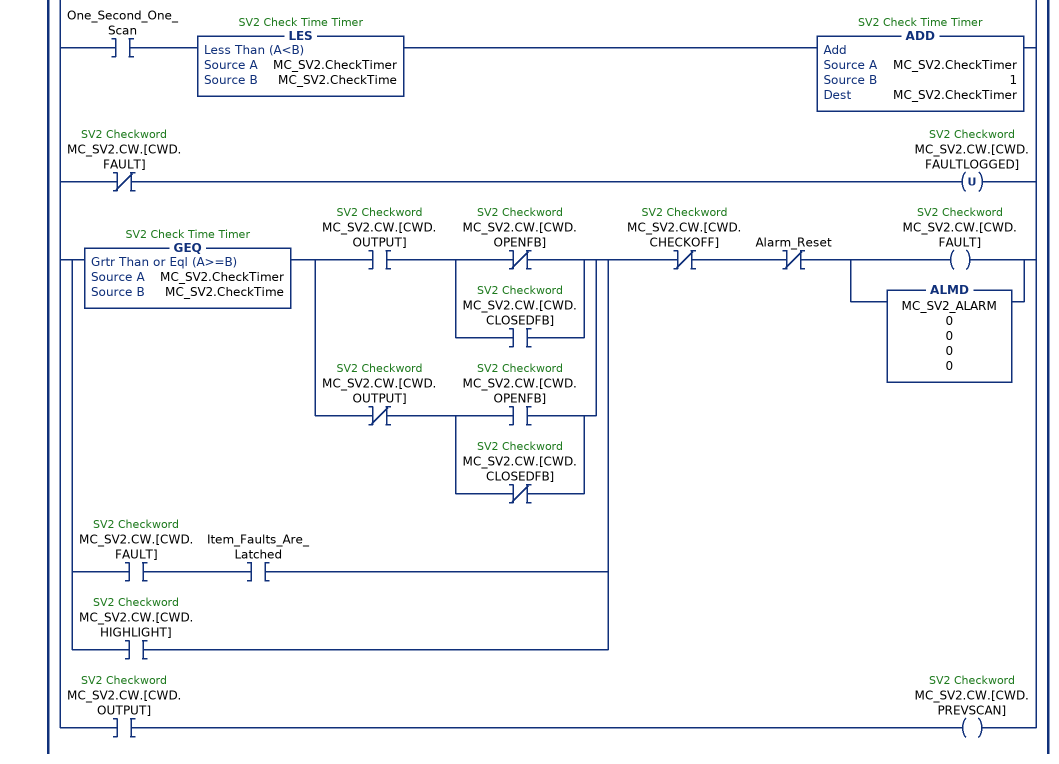
   46: [NEQ(MC_SV2.DriveBits,0) OTE(MC_SV2.CW.[CWD.AUTODRV]) ,[XIC(MC_SV2.CW.[CWD.AUTODRV]) XIO(MC_SV2.CW.[CWD.MANUAL]) ,XIC(MC_SV2.CW.[CWD.MANDRV]) XIC(MC_SV2.CW.[CWD.MANUAL]) ] OTE(MC_SV2.CW.[CWD.OUTPUT]) ,XIC(MC_SV2.CW.[CWD.OUTPUT]) OTE(MC_SV2_DR) ,XIC(S:FS) [OTU(MC_SV2.CW.[CWD.MANUAL]) ,LEQ(MC_SV2.CheckTime,0) MOV(Default_Check_Time,MC_SV2.CheckTime) ] ,[[XIC(MC_SV2_O) XIO(Item_Simulation_Flag) ,XIC(Item_Simulation_Flag) XIC(MC_SV2.CW.[CWD.OUTPUT]) XIO(MC_SV2.CW.[CWD.SIMFAIL]) ] OTE(MC_SV2.CW.[CWD.OPENFB]) ,[XIC(MC_SV2_C) XIO(Item_Simulation_Flag) ,XIC(Item_Simulation_Flag) XIO(MC_SV2.CW.[CWD.OUTPUT]) XIO(MC_SV2.CW.[CWD.SIMFAIL]) ] OTE(MC_SV2.CW.[CWD.CLOSEDFB]) ] ,[XIC(MC_SV2.CW.[CWD.OUTPUT]) XIO(MC_SV2.CW.[CWD.PREVSCAN]) ,XIO(MC_SV2.CW.[CWD.OUTPUT]) XIC(MC_SV2.CW.[CWD.PREVSCAN]) ] CLR(MC_SV2.CheckTimer) ,XIC(One_Second_One_Scan) LES(MC_SV2.CheckTimer,MC_SV2.CheckTime) ADD(MC_SV2.CheckTimer,1,MC_SV2.CheckTimer) ,XIO(MC_SV2.CW.[CWD.FAULT]) OTU(MC_SV2.CW.[CWD.FAULTLOGGED]) ,[GEQ(MC_SV2.CheckTimer,MC_SV2.CheckTime) [XIC(MC_SV2.CW.[CWD.OUTPUT]) [XIO(MC_SV2.CW.[CWD.OPENFB]) ,XIC(MC_SV2.CW.[CWD.CLOSEDFB]) ] ,XIO(MC_SV2.CW.[CWD.OUTPUT]) [XIC(MC_SV2.CW.[CWD.OPENFB]) ,XIO(MC_SV2.CW.[CWD.CLOSEDFB]) ] ] ,XIC(MC_SV2.CW.[CWD.FAULT]) XIC(Item_Faults_Are_Latched) ,XIC(MC_SV2.CW.[CWD.HIGHLIGHT]) ] XIO(MC_SV2.CW.[CWD.CHECKOFF]) XIO(Alarm_Reset) [OTE(MC_SV2.CW.[CWD.FAULT]) ,ALMD(MC_SV2_ALARM,0,0,0,0) ] ,XIC(MC_SV2.CW.[CWD.OUTPUT]) OTE(MC_SV2.CW.[CWD.PREVSCAN]) ];
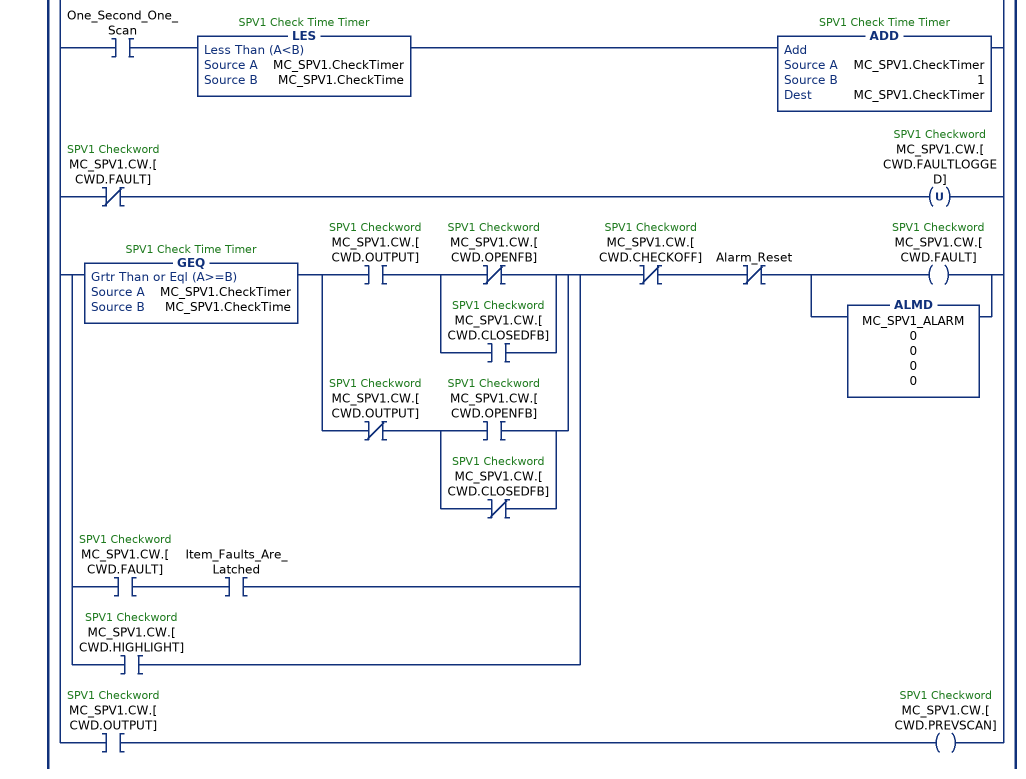
   47: [NEQ(MC_SPV1.DriveBits,0) OTE(MC_SPV1.CW.[CWD.AUTODRV]) ,[XIC(MC_SPV1.CW.[CWD.AUTODRV]) XIO(MC_SPV1.CW.[CWD.MANUAL]) ,XIC(MC_SPV1.CW.[CWD.MANDRV]) XIC(MC_SPV1.CW.[CWD.MANUAL]) ] OTE(MC_SPV1.CW.[CWD.OUTPUT]) ,XIC(MC_SPV1.CW.[CWD.OUTPUT]) OTE(MC_SPV1_DR) ,XIC(S:FS) [OTU(MC_SPV1.CW.[CWD.MANUAL]) ,LEQ(MC_SPV1.CheckTime,0) MOV(Default_Check_Time,MC_SPV1.CheckTime) ] ,[[XIC(MC_SPV1_O) XIO(Item_Simulation_Flag) ,XIC(Item_Simulation_Flag) XIC(MC_SPV1.CW.[CWD.OUTPUT]) XIO(MC_SPV1.CW.[CWD.SIMFAIL]) ] OTE(MC_SPV1.CW.[CWD.OPENFB]) ,[XIC(MC_SPV1_C) XIO(Item_Simulation_Flag) ,XIC(Item_Simulation_Flag) XIO(MC_SPV1.CW.[CWD.OUTPUT]) XIO(MC_SPV1.CW.[CWD.SIMFAIL]) ] OTE(MC_SPV1.CW.[CWD.CLOSEDFB]) ] ,[XIC(MC_SPV1.CW.[CWD.OUTPUT]) XIO(MC_SPV1.CW.[CWD.PREVSCAN]) ,XIO(MC_SPV1.CW.[CWD.OUTPUT]) XIC(MC_SPV1.CW.[CWD.PREVSCAN]) ] CLR(MC_SPV1.CheckTimer) ,XIC(One_Second_One_Scan) LES(MC_SPV1.CheckTimer,MC_SPV1.CheckTime) ADD(MC_SPV1.CheckTimer,1,MC_SPV1.CheckTimer) ,XIO(MC_SPV1.CW.[CWD.FAULT]) OTU(MC_SPV1.CW.[CWD.FAULTLOGGED]) ,[GEQ(MC_SPV1.CheckTimer,MC_SPV1.CheckTime) [XIC(MC_SPV1.CW.[CWD.OUTPUT]) [XIO(MC_SPV1.CW.[CWD.OPENFB]) ,XIC(MC_SPV1.CW.[CWD.CLOSEDFB]) ] ,XIO(MC_SPV1.CW.[CWD.OUTPUT]) [XIC(MC_SPV1.CW.[CWD.OPENFB]) ,XIO(MC_SPV1.CW.[CWD.CLOSEDFB]) ] ] ,XIC(MC_SPV1.CW.[CWD.FAULT]) XIC(Item_Faults_Are_Latched) ,XIC(MC_SPV1.CW.[CWD.HIGHLIGHT]) ] XIO(MC_SPV1.CW.[CWD.CHECKOFF]) XIO(Alarm_Reset) [OTE(MC_SPV1.CW.[CWD.FAULT]) ,ALMD(MC_SPV1_ALARM,0,0,0,0) ] ,XIC(MC_SPV1.CW.[CWD.OUTPUT]) OTE(MC_SPV1.CW.[CWD.PREVSCAN]) ];
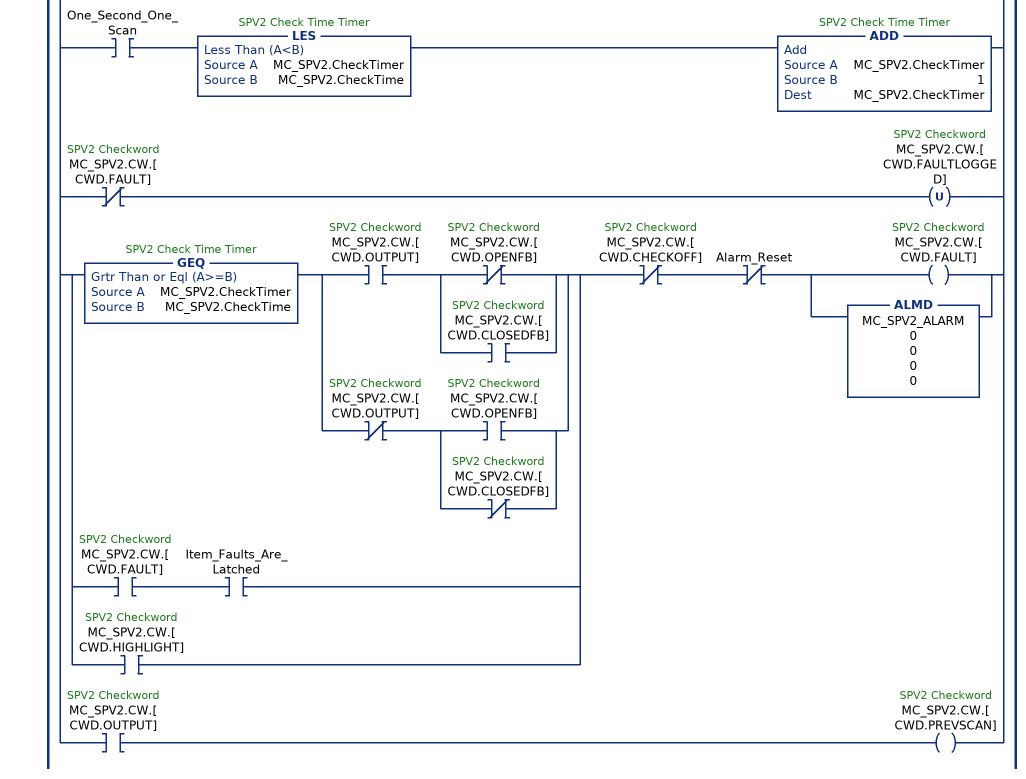
   48: [NEQ(MC_SPV2.DriveBits,0) OTE(MC_SPV2.CW.[CWD.AUTODRV]) ,[XIC(MC_SPV2.CW.[CWD.AUTODRV]) XIO(MC_SPV2.CW.[CWD.MANUAL]) ,XIC(MC_SPV2.CW.[CWD.MANDRV]) XIC(MC_SPV2.CW.[CWD.MANUAL]) ] OTE(MC_SPV2.CW.[CWD.OUTPUT]) ,XIC(MC_SPV2.CW.[CWD.OUTPUT]) OTE(MC_SPV2_DR) ,XIC(S:FS) [OTU(MC_SPV2.CW.[CWD.MANUAL]) ,LEQ(MC_SPV2.CheckTime,0) MOV(Default_Check_Time,MC_SPV2.CheckTime) ] ,[[XIC(MC_SPV2_O) XIO(Item_Simulation_Flag) ,XIC(Item_Simulation_Flag) XIC(MC_SPV2.CW.[CWD.OUTPUT]) XIO(MC_SPV2.CW.[CWD.SIMFAIL]) ] OTE(MC_SPV2.CW.[CWD.OPENFB]) ,[XIC(MC_SPV2_C) XIO(Item_Simulation_Flag) ,XIC(Item_Simulation_Flag) XIO(MC_SPV2.CW.[CWD.OUTPUT]) XIO(MC_SPV2.CW.[CWD.SIMFAIL]) ] OTE(MC_SPV2.CW.[CWD.CLOSEDFB]) ] ,[XIC(MC_SPV2.CW.[CWD.OUTPUT]) XIO(MC_SPV2.CW.[CWD.PREVSCAN]) ,XIO(MC_SPV2.CW.[CWD.OUTPUT]) XIC(MC_SPV2.CW.[CWD.PREVSCAN]) ] CLR(MC_SPV2.CheckTimer) ,XIC(One_Second_One_Scan) LES(MC_SPV2.CheckTimer,MC_SPV2.CheckTime) ADD(MC_SPV2.CheckTimer,1,MC_SPV2.CheckTimer) ,XIO(MC_SPV2.CW.[CWD.FAULT]) OTU(MC_SPV2.CW.[CWD.FAULTLOGGED]) ,[GEQ(MC_SPV2.CheckTimer,MC_SPV2.CheckTime) [XIC(MC_SPV2.CW.[CWD.OUTPUT]) [XIO(MC_SPV2.CW.[CWD.OPENFB]) ,XIC(MC_SPV2.CW.[CWD.CLOSEDFB]) ] ,XIO(MC_SPV2.CW.[CWD.OUTPUT]) [XIC(MC_SPV2.CW.[CWD.OPENFB]) ,XIO(MC_SPV2.CW.[CWD.CLOSEDFB]) ] ] ,XIC(MC_SPV2.CW.[CWD.FAULT]) XIC(Item_Faults_Are_Latched) ,XIC(MC_SPV2.CW.[CWD.HIGHLIGHT]) ] XIO(MC_SPV2.CW.[CWD.CHECKOFF]) XIO(Alarm_Reset) [OTE(MC_SPV2.CW.[CWD.FAULT]) ,ALMD(MC_SPV2_ALARM,0,0,0,0) ] ,XIC(MC_SPV2.CW.[CWD.OUTPUT]) OTE(MC_SPV2.CW.[CWD.PREVSCAN]) ];
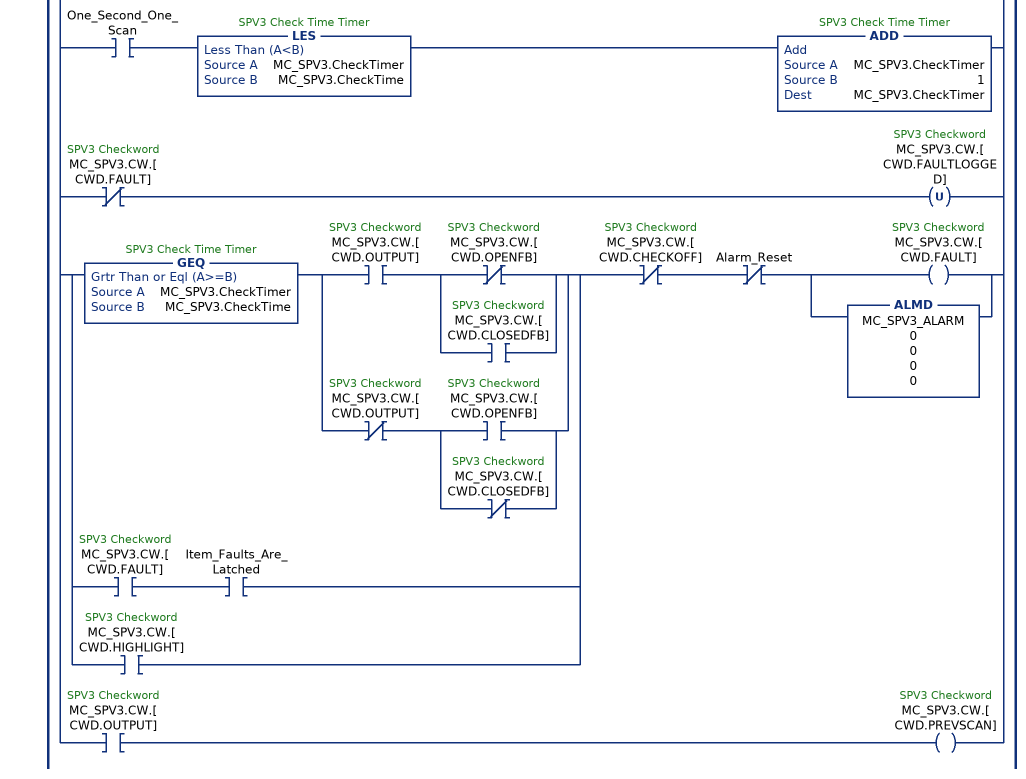
   49: [NEQ(MC_SPV3.DriveBits,0) OTE(MC_SPV3.CW.[CWD.AUTODRV]) ,[XIC(MC_SPV3.CW.[CWD.AUTODRV]) XIO(MC_SPV3.CW.[CWD.MANUAL]) ,XIC(MC_SPV3.CW.[CWD.MANDRV]) XIC(MC_SPV3.CW.[CWD.MANUAL]) ] OTE(MC_SPV3.CW.[CWD.OUTPUT]) ,XIC(MC_SPV3.CW.[CWD.OUTPUT]) OTE(MC_SPV3_DR) ,XIC(S:FS) [OTU(MC_SPV3.CW.[CWD.MANUAL]) ,LEQ(MC_SPV3.CheckTime,0) MOV(Default_Check_Time,MC_SPV3.CheckTime) ] ,[[XIC(MC_SPV3_O) XIO(Item_Simulation_Flag) ,XIC(Item_Simulation_Flag) XIC(MC_SPV3.CW.[CWD.OUTPUT]) XIO(MC_SPV3.CW.[CWD.SIMFAIL]) ] OTE(MC_SPV3.CW.[CWD.OPENFB]) ,[XIC(MC_SPV3_C) XIO(Item_Simulation_Flag) ,XIC(Item_Simulation_Flag) XIO(MC_SPV3.CW.[CWD.OUTPUT]) XIO(MC_SPV3.CW.[CWD.SIMFAIL]) ] OTE(MC_SPV3.CW.[CWD.CLOSEDFB]) ] ,[XIC(MC_SPV3.CW.[CWD.OUTPUT]) XIO(MC_SPV3.CW.[CWD.PREVSCAN]) ,XIO(MC_SPV3.CW.[CWD.OUTPUT]) XIC(MC_SPV3.CW.[CWD.PREVSCAN]) ] CLR(MC_SPV3.CheckTimer) ,XIC(One_Second_One_Scan) LES(MC_SPV3.CheckTimer,MC_SPV3.CheckTime) ADD(MC_SPV3.CheckTimer,1,MC_SPV3.CheckTimer) ,XIO(MC_SPV3.CW.[CWD.FAULT]) OTU(MC_SPV3.CW.[CWD.FAULTLOGGED]) ,[GEQ(MC_SPV3.CheckTimer,MC_SPV3.CheckTime) [XIC(MC_SPV3.CW.[CWD.OUTPUT]) [XIO(MC_SPV3.CW.[CWD.OPENFB]) ,XIC(MC_SPV3.CW.[CWD.CLOSEDFB]) ] ,XIO(MC_SPV3.CW.[CWD.OUTPUT]) [XIC(MC_SPV3.CW.[CWD.OPENFB]) ,XIO(MC_SPV3.CW.[CWD.CLOSEDFB]) ] ] ,XIC(MC_SPV3.CW.[CWD.FAULT]) XIC(Item_Faults_Are_Latched) ,XIC(MC_SPV3.CW.[CWD.HIGHLIGHT]) ] XIO(MC_SPV3.CW.[CWD.CHECKOFF]) XIO(Alarm_Reset) [OTE(MC_SPV3.CW.[CWD.FAULT]) ,ALMD(MC_SPV3_ALARM,0,0,0,0) ] ,XIC(MC_SPV3.CW.[CWD.OUTPUT]) OTE(MC_SPV3.CW.[CWD.PREVSCAN]) ];
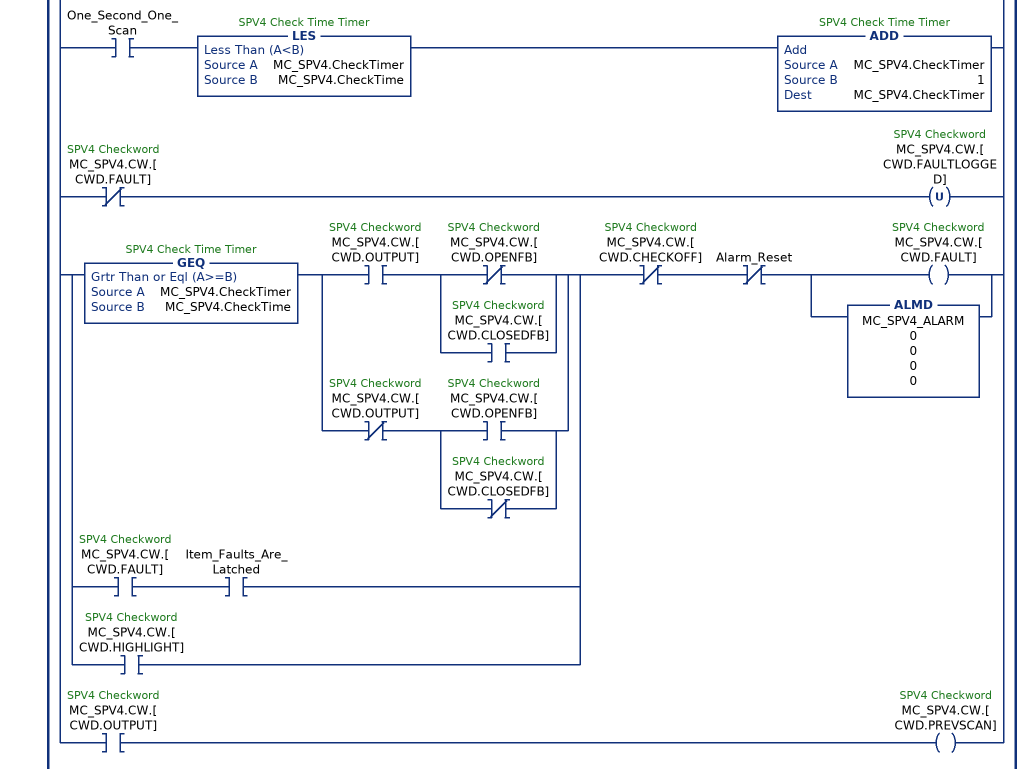
   50: [NEQ(MC_SPV4.DriveBits,0) OTE(MC_SPV4.CW.[CWD.AUTODRV]) ,[XIC(MC_SPV4.CW.[CWD.AUTODRV]) XIO(MC_SPV4.CW.[CWD.MANUAL]) ,XIC(MC_SPV4.CW.[CWD.MANDRV]) XIC(MC_SPV4.CW.[CWD.MANUAL]) ] OTE(MC_SPV4.CW.[CWD.OUTPUT]) ,XIC(MC_SPV4.CW.[CWD.OUTPUT]) OTE(MC_SPV4_DR) ,XIC(S:FS) [OTU(MC_SPV4.CW.[CWD.MANUAL]) ,LEQ(MC_SPV4.CheckTime,0) MOV(Default_Check_Time,MC_SPV4.CheckTime) ] ,[[XIC(MC_SPV4_O) XIO(Item_Simulation_Flag) ,XIC(Item_Simulation_Flag) XIC(MC_SPV4.CW.[CWD.OUTPUT]) XIO(MC_SPV4.CW.[CWD.SIMFAIL]) ] OTE(MC_SPV4.CW.[CWD.OPENFB]) ,[XIC(MC_SPV4_C) XIO(Item_Simulation_Flag) ,XIC(Item_Simulation_Flag) XIO(MC_SPV4.CW.[CWD.OUTPUT]) XIO(MC_SPV4.CW.[CWD.SIMFAIL]) ] OTE(MC_SPV4.CW.[CWD.CLOSEDFB]) ] ,[XIC(MC_SPV4.CW.[CWD.OUTPUT]) XIO(MC_SPV4.CW.[CWD.PREVSCAN]) ,XIO(MC_SPV4.CW.[CWD.OUTPUT]) XIC(MC_SPV4.CW.[CWD.PREVSCAN]) ] CLR(MC_SPV4.CheckTimer) ,XIC(One_Second_One_Scan) LES(MC_SPV4.CheckTimer,MC_SPV4.CheckTime) ADD(MC_SPV4.CheckTimer,1,MC_SPV4.CheckTimer) ,XIO(MC_SPV4.CW.[CWD.FAULT]) OTU(MC_SPV4.CW.[CWD.FAULTLOGGED]) ,[GEQ(MC_SPV4.CheckTimer,MC_SPV4.CheckTime) [XIC(MC_SPV4.CW.[CWD.OUTPUT]) [XIO(MC_SPV4.CW.[CWD.OPENFB]) ,XIC(MC_SPV4.CW.[CWD.CLOSEDFB]) ] ,XIO(MC_SPV4.CW.[CWD.OUTPUT]) [XIC(MC_SPV4.CW.[CWD.OPENFB]) ,XIO(MC_SPV4.CW.[CWD.CLOSEDFB]) ] ] ,XIC(MC_SPV4.CW.[CWD.FAULT]) XIC(Item_Faults_Are_Latched) ,XIC(MC_SPV4.CW.[CWD.HIGHLIGHT]) ] XIO(MC_SPV4.CW.[CWD.CHECKOFF]) XIO(Alarm_Reset) [OTE(MC_SPV4.CW.[CWD.FAULT]) ,ALMD(MC_SPV4_ALARM,0,0,0,0) ] ,XIC(MC_SPV4.CW.[CWD.OUTPUT]) OTE(MC_SPV4.CW.[CWD.PREVSCAN]) ];
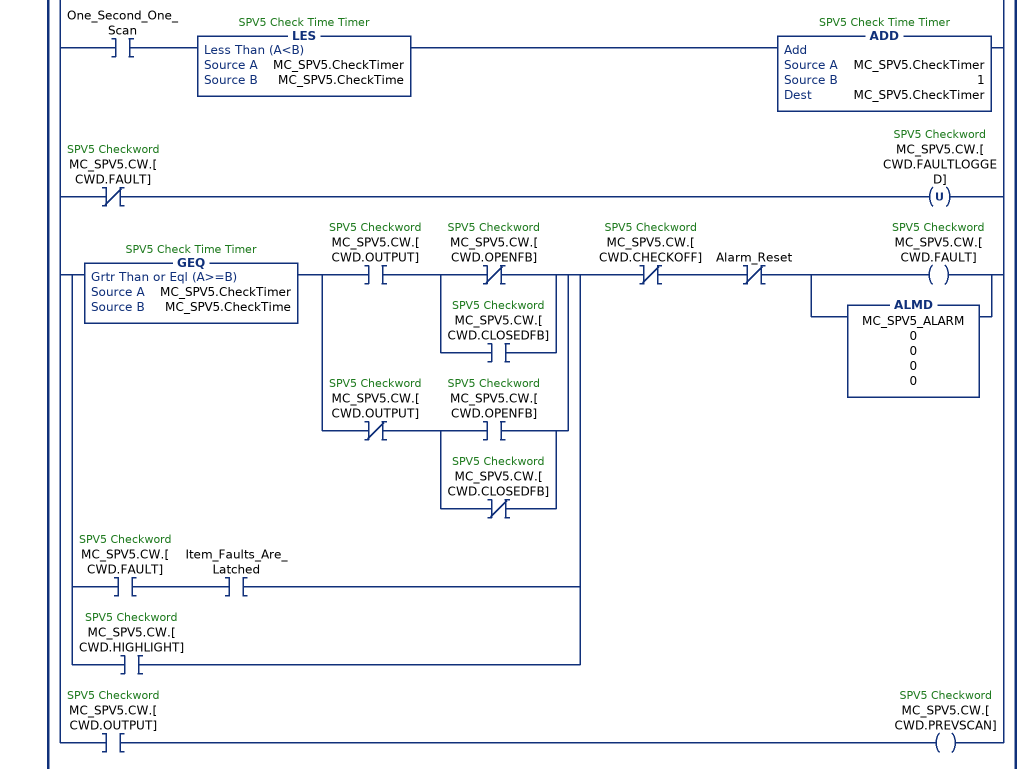
   51: [NEQ(MC_SPV5.DriveBits,0) OTE(MC_SPV5.CW.[CWD.AUTODRV]) ,[XIC(MC_SPV5.CW.[CWD.AUTODRV]) XIO(MC_SPV5.CW.[CWD.MANUAL]) ,XIC(MC_SPV5.CW.[CWD.MANDRV]) XIC(MC_SPV5.CW.[CWD.MANUAL]) ] OTE(MC_SPV5.CW.[CWD.OUTPUT]) ,XIC(MC_SPV5.CW.[CWD.OUTPUT]) OTE(MC_SPV5_DR) ,XIC(S:FS) [OTU(MC_SPV5.CW.[CWD.MANUAL]) ,LEQ(MC_SPV5.CheckTime,0) MOV(Default_Check_Time,MC_SPV5.CheckTime) ] ,[[XIC(MC_SPV5_O) XIO(Item_Simulation_Flag) ,XIC(Item_Simulation_Flag) XIC(MC_SPV5.CW.[CWD.OUTPUT]) XIO(MC_SPV5.CW.[CWD.SIMFAIL]) ] OTE(MC_SPV5.CW.[CWD.OPENFB]) ,[XIC(MC_SPV5_C) XIO(Item_Simulation_Flag) ,XIC(Item_Simulation_Flag) XIO(MC_SPV5.CW.[CWD.OUTPUT]) XIO(MC_SPV5.CW.[CWD.SIMFAIL]) ] OTE(MC_SPV5.CW.[CWD.CLOSEDFB]) ] ,[XIC(MC_SPV5.CW.[CWD.OUTPUT]) XIO(MC_SPV5.CW.[CWD.PREVSCAN]) ,XIO(MC_SPV5.CW.[CWD.OUTPUT]) XIC(MC_SPV5.CW.[CWD.PREVSCAN]) ] CLR(MC_SPV5.CheckTimer) ,XIC(One_Second_One_Scan) LES(MC_SPV5.CheckTimer,MC_SPV5.CheckTime) ADD(MC_SPV5.CheckTimer,1,MC_SPV5.CheckTimer) ,XIO(MC_SPV5.CW.[CWD.FAULT]) OTU(MC_SPV5.CW.[CWD.FAULTLOGGED]) ,[GEQ(MC_SPV5.CheckTimer,MC_SPV5.CheckTime) [XIC(MC_SPV5.CW.[CWD.OUTPUT]) [XIO(MC_SPV5.CW.[CWD.OPENFB]) ,XIC(MC_SPV5.CW.[CWD.CLOSEDFB]) ] ,XIO(MC_SPV5.CW.[CWD.OUTPUT]) [XIC(MC_SPV5.CW.[CWD.OPENFB]) ,XIO(MC_SPV5.CW.[CWD.CLOSEDFB]) ] ] ,XIC(MC_SPV5.CW.[CWD.FAULT]) XIC(Item_Faults_Are_Latched) ,XIC(MC_SPV5.CW.[CWD.HIGHLIGHT]) ] XIO(MC_SPV5.CW.[CWD.CHECKOFF]) XIO(Alarm_Reset) [OTE(MC_SPV5.CW.[CWD.FAULT]) ,ALMD(MC_SPV5_ALARM,0,0,0,0) ] ,XIC(MC_SPV5.CW.[CWD.OUTPUT]) OTE(MC_SPV5.CW.[CWD.PREVSCAN]) ];
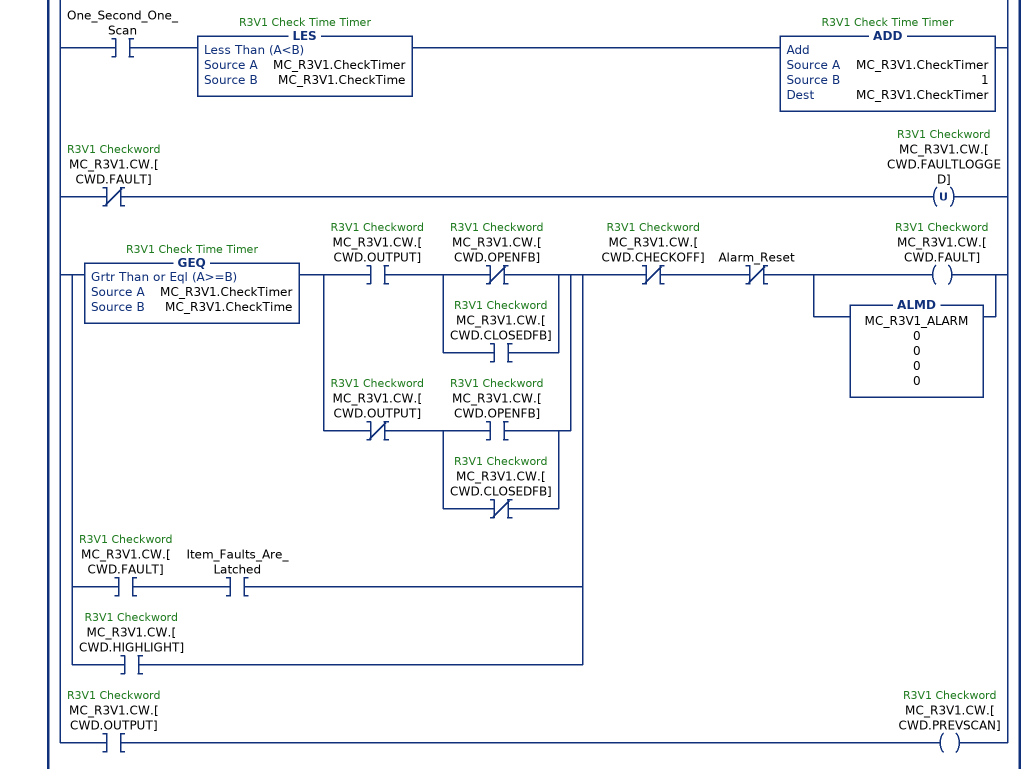
   52: [NEQ(MC_R3V1.DriveBits,0) OTE(MC_R3V1.CW.[CWD.AUTODRV]) ,[XIC(MC_R3V1.CW.[CWD.AUTODRV]) XIO(MC_R3V1.CW.[CWD.MANUAL]) ,XIC(MC_R3V1.CW.[CWD.MANDRV]) XIC(MC_R3V1.CW.[CWD.MANUAL]) ] OTE(MC_R3V1.CW.[CWD.OUTPUT]) ,XIC(MC_R3V1.CW.[CWD.OUTPUT]) OTE(MC_R3V1_DR) ,XIC(S:FS) [OTU(MC_R3V1.CW.[CWD.MANUAL]) ,LEQ(MC_R3V1.CheckTime,0) MOV(Default_Check_Time,MC_R3V1.CheckTime) ] ,[[XIC(MC_R3V1_O) XIO(Item_Simulation_Flag) ,XIC(Item_Simulation_Flag) XIC(MC_R3V1.CW.[CWD.OUTPUT]) XIO(MC_R3V1.CW.[CWD.SIMFAIL]) ] OTE(MC_R3V1.CW.[CWD.OPENFB]) ,[XIC(MC_R3V1_C) XIO(Item_Simulation_Flag) ,XIC(Item_Simulation_Flag) XIO(MC_R3V1.CW.[CWD.OUTPUT]) XIO(MC_R3V1.CW.[CWD.SIMFAIL]) ] OTE(MC_R3V1.CW.[CWD.CLOSEDFB]) ] ,[XIC(MC_R3V1.CW.[CWD.OUTPUT]) XIO(MC_R3V1.CW.[CWD.PREVSCAN]) ,XIO(MC_R3V1.CW.[CWD.OUTPUT]) XIC(MC_R3V1.CW.[CWD.PREVSCAN]) ] CLR(MC_R3V1.CheckTimer) ,XIC(One_Second_One_Scan) LES(MC_R3V1.CheckTimer,MC_R3V1.CheckTime) ADD(MC_R3V1.CheckTimer,1,MC_R3V1.CheckTimer) ,XIO(MC_R3V1.CW.[CWD.FAULT]) OTU(MC_R3V1.CW.[CWD.FAULTLOGGED]) ,[GEQ(MC_R3V1.CheckTimer,MC_R3V1.CheckTime) [XIC(MC_R3V1.CW.[CWD.OUTPUT]) [XIO(MC_R3V1.CW.[CWD.OPENFB]) ,XIC(MC_R3V1.CW.[CWD.CLOSEDFB]) ] ,XIO(MC_R3V1.CW.[CWD.OUTPUT]) [XIC(MC_R3V1.CW.[CWD.OPENFB]) ,XIO(MC_R3V1.CW.[CWD.CLOSEDFB]) ] ] ,XIC(MC_R3V1.CW.[CWD.FAULT]) XIC(Item_Faults_Are_Latched) ,XIC(MC_R3V1.CW.[CWD.HIGHLIGHT]) ] XIO(MC_R3V1.CW.[CWD.CHECKOFF]) XIO(Alarm_Reset) [OTE(MC_R3V1.CW.[CWD.FAULT]) ,ALMD(MC_R3V1_ALARM,0,0,0,0) ] ,XIC(MC_R3V1.CW.[CWD.OUTPUT]) OTE(MC_R3V1.CW.[CWD.PREVSCAN]) ];
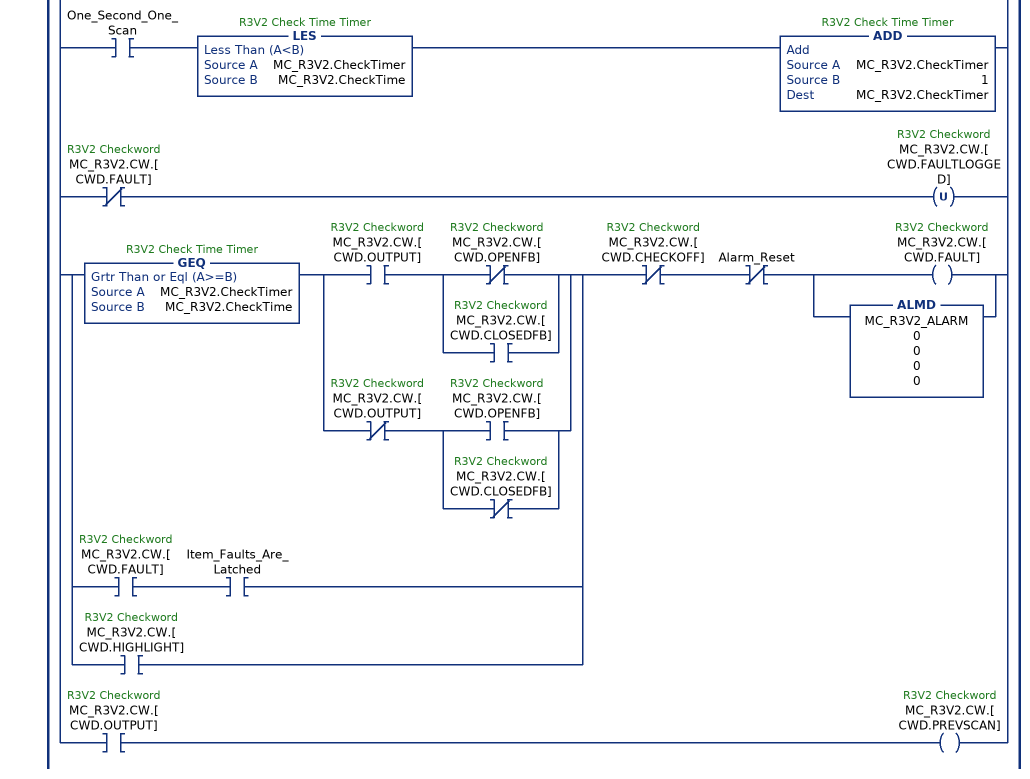
   53: [NEQ(MC_R3V2.DriveBits,0) OTE(MC_R3V2.CW.[CWD.AUTODRV]) ,[XIC(MC_R3V2.CW.[CWD.AUTODRV]) XIO(MC_R3V2.CW.[CWD.MANUAL]) ,XIC(MC_R3V2.CW.[CWD.MANDRV]) XIC(MC_R3V2.CW.[CWD.MANUAL]) ] OTE(MC_R3V2.CW.[CWD.OUTPUT]) ,XIC(MC_R3V2.CW.[CWD.OUTPUT]) OTE(MC_R3V2_DR) ,XIC(S:FS) [OTU(MC_R3V2.CW.[CWD.MANUAL]) ,LEQ(MC_R3V2.CheckTime,0) MOV(Default_Check_Time,MC_R3V2.CheckTime) ] ,[[XIC(MC_R3V2_O) XIO(Item_Simulation_Flag) ,XIC(Item_Simulation_Flag) XIC(MC_R3V2.CW.[CWD.OUTPUT]) XIO(MC_R3V2.CW.[CWD.SIMFAIL]) ] OTE(MC_R3V2.CW.[CWD.OPENFB]) ,[XIC(MC_R3V2_C) XIO(Item_Simulation_Flag) ,XIC(Item_Simulation_Flag) XIO(MC_R3V2.CW.[CWD.OUTPUT]) XIO(MC_R3V2.CW.[CWD.SIMFAIL]) ] OTE(MC_R3V2.CW.[CWD.CLOSEDFB]) ] ,[XIC(MC_R3V2.CW.[CWD.OUTPUT]) XIO(MC_R3V2.CW.[CWD.PREVSCAN]) ,XIO(MC_R3V2.CW.[CWD.OUTPUT]) XIC(MC_R3V2.CW.[CWD.PREVSCAN]) ] CLR(MC_R3V2.CheckTimer) ,XIC(One_Second_One_Scan) LES(MC_R3V2.CheckTimer,MC_R3V2.CheckTime) ADD(MC_R3V2.CheckTimer,1,MC_R3V2.CheckTimer) ,XIO(MC_R3V2.CW.[CWD.FAULT]) OTU(MC_R3V2.CW.[CWD.FAULTLOGGED]) ,[GEQ(MC_R3V2.CheckTimer,MC_R3V2.CheckTime) [XIC(MC_R3V2.CW.[CWD.OUTPUT]) [XIO(MC_R3V2.CW.[CWD.OPENFB]) ,XIC(MC_R3V2.CW.[CWD.CLOSEDFB]) ] ,XIO(MC_R3V2.CW.[CWD.OUTPUT]) [XIC(MC_R3V2.CW.[CWD.OPENFB]) ,XIO(MC_R3V2.CW.[CWD.CLOSEDFB]) ] ] ,XIC(MC_R3V2.CW.[CWD.FAULT]) XIC(Item_Faults_Are_Latched) ,XIC(MC_R3V2.CW.[CWD.HIGHLIGHT]) ] XIO(MC_R3V2.CW.[CWD.CHECKOFF]) XIO(Alarm_Reset) [OTE(MC_R3V2.CW.[CWD.FAULT]) ,ALMD(MC_R3V2_ALARM,0,0,0,0) ] ,XIC(MC_R3V2.CW.[CWD.OUTPUT]) OTE(MC_R3V2.CW.[CWD.PREVSCAN]) ];
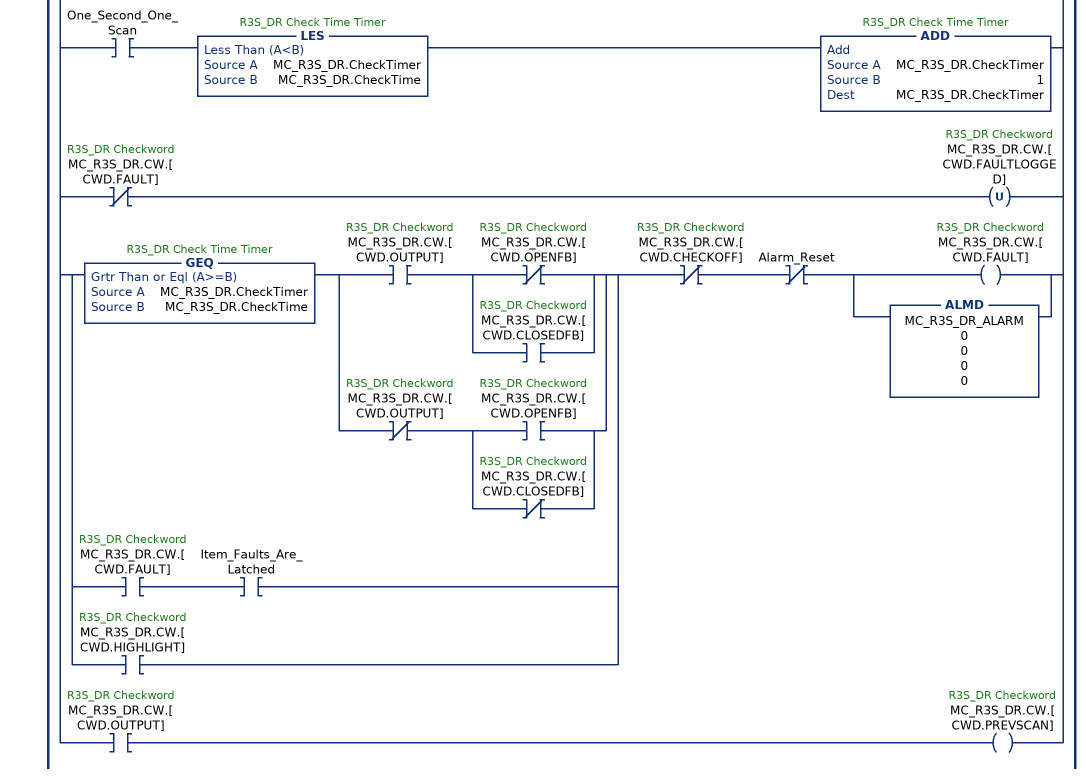
   54: [NEQ(MC_R3S_DR.DriveBits,0) OTE(MC_R3S_DR.CW.[CWD.AUTODRV]) ,[XIC(MC_R3S_DR.CW.[CWD.AUTODRV]) XIO(MC_R3S_DR.CW.[CWD.MANUAL]) ,XIC(MC_R3S_DR.CW.[CWD.MANDRV]) XIC(MC_R3S_DR.CW.[CWD.MANUAL]) ] OTE(MC_R3S_DR.CW.[CWD.OUTPUT]) ,XIC(MC_R3S_DR.CW.[CWD.OUTPUT]) OTE(MC_R3S_DR_DR) ,XIC(S:FS) [OTU(MC_R3S_DR.CW.[CWD.MANUAL]) ,LEQ(MC_R3S_DR.CheckTime,0) MOV(Default_Check_Time,MC_R3S_DR.CheckTime) ] ,[[XIC(MC_R3S_DR_O) XIO(Item_Simulation_Flag) ,XIC(Item_Simulation_Flag) XIC(MC_R3S_DR.CW.[CWD.OUTPUT]) XIO(MC_R3S_DR.CW.[CWD.SIMFAIL]) ] OTE(MC_R3S_DR.CW.[CWD.OPENFB]) ,[XIC(MC_R3S_DR_C) XIO(Item_Simulation_Flag) ,XIC(Item_Simulation_Flag) XIO(MC_R3S_DR.CW.[CWD.OUTPUT]) XIO(MC_R3S_DR.CW.[CWD.SIMFAIL]) ] OTE(MC_R3S_DR.CW.[CWD.CLOSEDFB]) ] ,[XIC(MC_R3S_DR.CW.[CWD.OUTPUT]) XIO(MC_R3S_DR.CW.[CWD.PREVSCAN]) ,XIO(MC_R3S_DR.CW.[CWD.OUTPUT]) XIC(MC_R3S_DR.CW.[CWD.PREVSCAN]) ] CLR(MC_R3S_DR.CheckTimer) ,XIC(One_Second_One_Scan) LES(MC_R3S_DR.CheckTimer,MC_R3S_DR.CheckTime) ADD(MC_R3S_DR.CheckTimer,1,MC_R3S_DR.CheckTimer) ,XIO(MC_R3S_DR.CW.[CWD.FAULT]) OTU(MC_R3S_DR.CW.[CWD.FAULTLOGGED]) ,[GEQ(MC_R3S_DR.CheckTimer,MC_R3S_DR.CheckTime) [XIC(MC_R3S_DR.CW.[CWD.OUTPUT]) [XIO(MC_R3S_DR.CW.[CWD.OPENFB]) ,XIC(MC_R3S_DR.CW.[CWD.CLOSEDFB]) ] ,XIO(MC_R3S_DR.CW.[CWD.OUTPUT]) [XIC(MC_R3S_DR.CW.[CWD.OPENFB]) ,XIO(MC_R3S_DR.CW.[CWD.CLOSEDFB]) ] ] ,XIC(MC_R3S_DR.CW.[CWD.FAULT]) XIC(Item_Faults_Are_Latched) ,XIC(MC_R3S_DR.CW.[CWD.HIGHLIGHT]) ] XIO(MC_R3S_DR.CW.[CWD.CHECKOFF]) XIO(Alarm_Reset) [OTE(MC_R3S_DR.CW.[CWD.FAULT]) ,ALMD(MC_R3S_DR_ALARM,0,0,0,0) ] ,XIC(MC_R3S_DR.CW.[CWD.OUTPUT]) OTE(MC_R3S_DR.CW.[CWD.PREVSCAN]) ];
